               "DB919_ShotResultMach".ShotResult_Ma[1].Component.Comp[#Component].MaterialConsumption :=
               #TempConsumption +
               ("DB919_ShotResultMach".ShotResult_Ma[1].Component.Comp[#Component].Flow *
               "DB704_MH_Value".Mixinghead[#MHNumber].Corrvalue);

           ELSE
               "DB919_ShotResultMach".ShotResult_Ma[1].Component.Comp[#Component].MaterialConsumption :=
               #TempConsumption;

           END_IF;

       END_IF;
   END_FOR;
END_FUNCTION

ORGANIZATION_BLOCK "Cycle Execution"   // OB1, STL, ProgramCycle
TITLE = "Main Program Sweep (Cycle)"
{ S7_Optimized_Access := 'FALSE' }
VERSION : 0.1
   VAR_TEMP
      OB1_EV_CLASS : Byte;   // Bits 0-3 = 1 (Coming event), Bits 4-7 = 1 (Event class 1)
      OB1_SCAN_1 : Byte;   // 1 (Cold restart scan 1 of OB 1), 3 (Scan 2-n of OB 1)
      OB1_PRIORITY : Byte;   // Priority of OB Execution
      OB1_OB_NUMBR : Byte;   // 1 (Organization block 1, OB1)
      OB1_RESERVED_1 : Byte;   // Reserved for system
      OB1_RESERVED_2 : Byte;   // Reserved for system
      OB1_PREV_CYCLE : Int;   // Cycle time of previous OB1 scan (milliseconds)
      OB1_MIN_CYCLE : Int;   // Minimum cycle time of OB1 (milliseconds)
      OB1_MAX_CYCLE : Int;   // Maximum cycle time of OB1 (milliseconds)
      OB1_DATE_TIME : Date_And_Time;   // Date and time OB1 started
      Ret_Val_SFC51 : Int;
      SLZ_Header : Struct
         LENTHDR : Word;
         N_DR : Word;
      END_STRUCT;
      TmpMachineNo : Int;
      DPDPoff : Bool;
      RetValSFC : Int;
      DPDPon : Bool;
      D_ACT_DP_Busy : Bool;
   END_VAR
BEGIN

REGION Network 1: First PLC cycle
         A(;
         L     #OB1_SCAN_1;
         L     1;
         ==I;
         );
         =     "Flag_Erster_SPS_Zyklus";

   // --- Activate addresses of IO interface ProCan
         A     "Flag_Erster_SPS_Zyklus";
         S     "M1200_ActivateAdrProCan";
END_REGION

REGION Network 2: ProNet-Functions
         A     "Flag_Erster_SPS_Zyklus";
         R     "Flag_ToggleForDatarequest";

         CALL  "PNC_AI"
         ( RequestAll        := "Flag_Erster_SPS_Zyklus",
           AcknowledgeFaults := "DB009_Faults".Faults_Reset_FKT_M1,
           GOON              := "Flag_ToggleForDatarequest"
         );

         CALL  "PNC_Mixinghead"
         ( RequestAll        := "Flag_Erster_SPS_Zyklus",
           AcknowledgeFaults := "DB009_Faults".Faults_Reset_FKT_M1,
           GOON              := "Flag_ToggleForDatarequest"
         );

         CALL  "PNC_Flow"
         ( RequestAll        := "Flag_Erster_SPS_Zyklus",
           AcknowledgeFaults := "DB009_Faults".Faults_Reset_FKT_M1,
           GOON              := "Flag_ToggleForDatarequest"
         );

         AN    "Flag_ToggleForDatarequest";
         =     "Flag_ToggleForDatarequest";
END_REGION

REGION Network 3: Brücken für Inbetriebnahme
         CLR;
         =     "With_MC03";
         =     "With_MC04";
END_REGION

REGION Network 4: Handling Mould Editor
         CALL  "FB_MouldEditor_HMI", "FB_MouldEditor_HMI_DB"
         ( INiAmountMeteringUnits := "DB790_PlantParameter".AmountMeteringUnits,
           IOuMouldEditor_HMI     := "DB_MouldEditor_HMI".uData
         );
END_REGION

REGION Network 5: Analyse der Profinet- und Profibusbusteilnehmer
   // PN devices analyze
         CALL  DeviceStates
         ( LADDR   := "PN_Devices".LADDR,
           MODE    := "PN_Devices".MODE,
           Ret_Val := "PN_Devices".RETVAL,
           STATE   := "PN_Devices".Device_available
         );

   // PB devices analyze
         CALL  DeviceStates
         ( LADDR   := "PB_Devices".LADDR,
           MODE    := "PB_Devices".MODE,
           Ret_Val := "PB_Devices".RETVAL,
           STATE   := "PB_Devices".Device_available
         );
END_REGION

REGION Network 6: Tempering
   // Test
         CALL  "Baustein_1";

         O     "DB702_Tank_Value".Tank[1].With_Tempering_TempGeraet;
         O     "DB702_Tank_Value".Tank[1].With_Tempering_VKaltwasser;
         O     "DB702_Tank_Value".Tank[1].With_Tempering_Heizung;
         O     "DB702_Tank_Value".Tank[1].With_Tempering_WTRL;
         O     "DB702_Tank_Value".Tank[1].With_Tempering_WTmitFischer;
         O     "DB702_Tank_Value".Tank[1].With_Tempering_WTBypass;
         O     "DB702_Tank_Value".Tank[1].With_Tempering_WTVL;
   // Damit der Schalter für die Temperierung angezeigt wird
         =     "DB702_Tank_Value".Tank[1].With_Tempering;

         O     "DB702_Tank_Value".Tank[2].With_Tempering_TempGeraet;
         O     "DB702_Tank_Value".Tank[2].With_Tempering_VKaltwasser;
         O     "DB702_Tank_Value".Tank[2].With_Tempering_Heizung;
         O     "DB702_Tank_Value".Tank[2].With_Tempering_WTRL;
         O     "DB702_Tank_Value".Tank[2].With_Tempering_WTmitFischer;
         O     "DB702_Tank_Value".Tank[2].With_Tempering_WTBypass;
         O     "DB702_Tank_Value".Tank[2].With_Tempering_WTVL;
         =     "DB702_Tank_Value".Tank[2].With_Tempering;

         O     "DB702_Tank_Value".Tank[3].With_Tempering_TempGeraet;
         O     "DB702_Tank_Value".Tank[3].With_Tempering_VKaltwasser;
         O     "DB702_Tank_Value".Tank[3].With_Tempering_Heizung;
         O     "DB702_Tank_Value".Tank[3].With_Tempering_WTRL;
         O     "DB702_Tank_Value".Tank[3].With_Tempering_WTmitFischer;
         O     "DB702_Tank_Value".Tank[3].With_Tempering_WTBypass;
         O     "DB702_Tank_Value".Tank[3].With_Tempering_WTVL;
         =     "DB702_Tank_Value".Tank[3].With_Tempering;

         O     "DB702_Tank_Value".Tank[4].With_Tempering_TempGeraet;
         O     "DB702_Tank_Value".Tank[4].With_Tempering_VKaltwasser;
         O     "DB702_Tank_Value".Tank[4].With_Tempering_Heizung;
         O     "DB702_Tank_Value".Tank[4].With_Tempering_WTRL;
         O     "DB702_Tank_Value".Tank[4].With_Tempering_WTmitFischer;
         O     "DB702_Tank_Value".Tank[4].With_Tempering_WTBypass;
         O     "DB702_Tank_Value".Tank[4].With_Tempering_WTVL;
         =     "DB702_Tank_Value".Tank[4].With_Tempering;
END_REGION

REGION Network 7: Inputs external plant
   // MC1
   //      CALL  DPRD_DAT
   //         LADDR   :="PN-PN-Coupler_PU_MC1~IN___8_Byte"
   //         RET_VAL :=#RetValSFC
   //         RECORD  :="DB005_RS<->Extern".MC_Interface[1].Data_from_MC
   // MC2
   //     CALL  DPRD_DAT
   //         LADDR   :="PN-PN-Coupler_PU_MC2~IN__16_Byte"
   //         RET_VAL :=#RetValSFC
   //         RECORD  :="DB005_RS<->Extern".MC_Interface[2].Data_from_MC
   // MC3
   //      CALL  DPRD_DAT
   //         LADDR   :="PN-PN-Coupler_PU_MC3~IN__16_Byte"
   //         RET_VAL :=#RetValSFC
   //         RECORD  :="DB005_RS<->Extern".MC_Interface[3].Data_from_MC

   // MC4
   //      CALL  DPRD_DAT
   //         LADDR   :="PN-PN-Coupler_PU_MC4~IN__16_Byte"
   //         RET_VAL :=#RetValSFC
   //         RECORD  :="DB005_RS<->Extern".MC_Interface[4].Data_from_MC
END_REGION

REGION Network 8: Force Inputs
   //      L     "Interface_Signals_From_KMI":P
   //      T     %DB5.DBW20
   //      L     "Tag_35":P
   //      T     "DB005_RS<->Extern".MC_Interface[1].FromMC.Temperature_Tool01
   //      L     "Tag_36":P
   //      T     "DB005_RS<->Extern".MC_Interface[1].FromMC.Temperature_Tool02
   //      L     "Tag_37":P
   //      T     "DB005_RS<->Extern".MC_Interface[1].FromMC.Spare_6
   //      L     "Tag_38":P
   //      T     "DB005_RS<->Extern".MC_Interface[1].FromMC.Spare_8

   //      L     "Tag_39":P
   //      T     %DB5.DBW40
   //      L     "Tag_40":P
   //      T     "DB005_RS<->Extern".MC_Interface[2].FromMC.Temperature_Tool01
   //      L     "Tag_41":P
   //      T     "DB005_RS<->Extern".MC_Interface[2].FromMC.Temperature_Tool02
   //      L     "Tag_42":P
   //      T     "DB005_RS<->Extern".MC_Interface[2].FromMC.Spare_6
   //      L     "Tag_43":P
   //      T     "DB005_RS<->Extern".MC_Interface[2].FromMC.Spare_8
END_REGION

REGION Network 9: Check Profnet Slaves
   //
         CALL  DeviceStates
         ( LADDR   := 257,
           MODE    := 4,
           Ret_Val := #Ret_Val_SFC51,
           STATE   := "PN_DeviceState".StatePN
         );
   //
END_REGION

REGION Network 10: Interface Visu
         CALL  "FC5011_InterfaceHydraulik"
         ( Enable := 1
         );

         CALL  "FC5012_InterfaceTank"
         ( Enable := 1
         );

         CALL  "FC5013_InterfaceMetering"
         ( Enable := 1
         );

         CALL  "FC5014_InterfaceMixinghead"
         ( Enable := 1
         );

         CALL  "FC5020_InterfaceConfig"
         ( Enable := 1
         );

         CALL  "FC5900_InterfaceRobots"
         ( Enable := 1
         );
END_REGION

REGION Network 11: Program blocks
   //
         UC    "FB009_Faults";

   // machine 1
         UC    "FB011_OP_CirceMode_M1";
         UC    "FB012_MH_Hydraulic_M1";
         UC    "FB014_MH_SWU_M1";
         UC    "FB015_MeteringPump_M1";
   //     UC    "FB016_MeteringPump_Heating_M1"
         UC    "FB019_FoamingCycle_M1";
         UC    "FB017_CPiston_M1";

   // common function blocks
         UC    "FB100_Common_Aggregates_General";
         UC    "FB101_Common_Aggregates_C1";
         UC    "FB102_Common_Aggregates_C2";

         UC    "FB110_Interface_Prog_M1";
   //      UC    "FB111_Inerting"

         UC    "FB120_ProcanIO_RW";
   //      UC    "FB130_Tempering"
   //      UC    "FB140_ConfProCan"

         UC    "FB916_PV_LimitControl";

         UC    "FB919_PV_SetValueFoaming";
         UC    "FB920_ShotResult";

         UC    "FB930_FoamingData";

   //      UC    "FB1900_IF_Robots"

         UC    "FB1025_Service";

         CALL  "FC14_TP_Shortcuts";

   // Interface
         CALL  "FC2001_KM_FRA";
END_REGION

REGION Network 12: General functions
END_REGION

REGION Network 13: Outputs external plant
   // MC1
   //    CALL  DPWR_DAT
   //         LADDR   :="PN-PN-Coupler_PU_MC1~OUT___8_Byte"
   //         RECORD  :="DB005_RS<->Extern".MC_Interface[1].Data_to_MC
   //         RET_VAL :=#RetValSFC
   // MC2
   //     CALL  DPWR_DAT
   //         LADDR   :="PN-PN-Coupler_PU_MC2~OUT__16_Byte"
   //         RECORD  :="DB005_RS<->Extern".MC_Interface[2].Data_to_MC
   //         RET_VAL :=#RetValSFC
   // MC3
   //      CALL  DPWR_DAT
   //         LADDR   :="PN-PN-Coupler_PU_MC3~OUT__16_Byte"
   //         RECORD  :="DB005_RS<->Extern".MC_Interface[3].Data_to_MC
   //         RET_VAL :=#RetValSFC
   // MC4
   //      CALL  DPWR_DAT
   //         LADDR   :="PN-PN-Coupler_PU_MC4~OUT__16_Byte"
   //         RECORD  :="DB005_RS<->Extern".MC_Interface[4].Data_to_MC
   //         RET_VAL :=#RetValSFC
END_REGION

REGION Network 14: AllocationList
         CALL  "FB1931_ToolAllocationList", "FB1931_ToolAllocationList_DB";
END_REGION

REGION Network 15: Oszi
         CALL  "FC025_Oszilloskop";
         CALL  "FC117_INT_Umwandler";
END_REGION

REGION Network 16: TurnTable
   //    UC    "FB1001_TT"
END_REGION

REGION Network 17: RFID

   //      CALL  "FC030_BalluffReader 1"
   //      CALL  "FC031_BalluffReader 2"
END_REGION

REGION Network 18: Traceability
         CALL  "FC1500_ShotDataToMC";
END_REGION

REGION Network 19: Date and time
         CALL  "FC2170_TimeHandle";
   //-----
END_REGION

REGION Network 20: Network connection flag
         A     "Flag_00_500_Hertz";
         =     "Flag_Network";
END_REGION

REGION Network 21: delay_timer
         A     "new_shift";
         L     s5t#60s;
         SD    "delay_timer";
         A     "delay_timer";
         R     "new_shift";

         AN    "new_shift";
         R     "flag_delay_check_path";
         L     s5t#20s;
         SD    "Timer_check_path";
         A     "Timer_check_path";
         S     "flag_delay_check_path";
         R     "delay_timer";
END_REGION

REGION Network 22: IBN
         A     "AlwaysFALSE";
         R     "AlwaysFALSE";
         AN    "AlwaysTRUE";
         S     "AlwaysTRUE";
END_REGION
END_ORGANIZATION_BLOCK

ORGANIZATION_BLOCK "CYC_INT5"   // OB35, STL, CyclicInterrupt
TITLE = "Cyclic Interrupt"
{ S7_Optimized_Access := 'FALSE' }
AUTHOR : KT242
VERSION : 0.1
   VAR_TEMP
      OB35_EV_CLASS : Byte;   // Bits 0-3 = 1 (Coming event), Bits 4-7 = 1 (Event class 1)
      OB35_STRT_INF : Byte;   // 16#36 (OB 35 has started)
      OB35_PRIORITY : Byte;   // Priority of OB Execution
      OB35_OB_NUMBR : Byte;   // 35 (Organization block 35, OB35)
      OB35_RESERVED_1 : Byte;   // Reserved for system
      OB35_RESERVED_2 : Byte;   // Reserved for system
      OB35_PHASE_OFFSET : Word;   // Phase offset (msec)
      OB35_RESERVED_3 : Int;   // Reserved for system
      OB35_EXC_FREQ : Int;   // Frequency of execution (msec)
      OB35_DATE_TIME : Date_And_Time;   // Date and time OB35 started
      Temp_MH_Temp_C1 : Int;
      Temp_MH_Temp_C2 : Int;
      Temp_MH_Pressure_C1 : Int;
      Temp_MH_Pressure_C2 : Int;
      DINT_dummy : Real;
      dummy : Bool;
      Tenmp_flow_comp1 : DInt;
      Tenmp_flow_comp2 : DInt;
      Temp_ShotTimeAct : DInt;
      TempDBNo : Word;
      TempDWNo : DInt;
      TempRetClock : Int;
      TempDateTime : Date_And_Time;
      TempWritePointer : Int;
      EXC_FREQ_HE : Int;   // Execution frequency of heat exchangers
      TempSWU_MH01 : Bool;
      TempSWU_MH02 : Bool;
      TempSWU_MH03 : Bool;
      TempSWU_MH04 : Bool;
      TempSWU_MH05 : Bool;
      TempSWU_MH06 : Bool;
      TempSWU_MH07 : Bool;
      TempSWU_MH08 : Bool;
      TempSWU_MH09 : Bool;
      TempSWU_MH10 : Bool;
      Temp_CompFlowReal : Real;
      Temp_STimeReal : Real;
      CompUsedForShot : Array[1..16] of Bool;
   END_VAR
BEGIN

REGION Network 1: Read PV flowrate and calc. consumption of components machine 1
         A     "DB619_State_MPart".Cycle[1].Shotrelease;
         FP    "FHF_ShotreleaseM1";
         JCN   f101;
         L     0.0;
         T     "AmountFlowValuesMa1C1";
         T     "AmountFlowValuesMa1C2";
         T     "AmountFlowValuesMa1C3";
         T     "AmountFlowValuesMa1C4";
         T     "AmountFlowValuesMa1C5";
         T     "AmountFlowValuesMa1C6";
         T     "AmountFlowValuesMa1C7";
         T     "AmountFlowValuesMa1C8";
         T     "AmountFlowValuesMa1C9";
         T     "AmountFlowValuesMa1C10";
         T     "AmountFlowValuesMa1C11";
         T     "AmountFlowValuesMa1C12";

         T     "TotalFlowShotC01";
         T     "TotalFlowShotC02";
         T     "TotalFlowShotC03";
         T     "TotalFlowShotC04";
         T     "TotalFlowShotC05";
         T     "TotalFlowShotC06";
         T     "TotalFlowShotC07";
         T     "TotalFlowShotC08";
         T     "TotalFlowShotC09";
         T     "TotalFlowShotC10";
         T     "TotalFlowShotC11";
         T     "TotalFlowShotC12";


         T     "DB919_ShotResultMach".ShotResult_Ma[1].General.FoamingTime;
         T     "DB919_ShotResultMach".ShotResult_Ma[1].Component.Comp[1].Flow;
         T     "DB919_ShotResultMach".ShotResult_Ma[1].Component.Comp[2].Flow;
         T     "DB919_ShotResultMach".ShotResult_Ma[1].Component.Comp[3].Flow;
         T     "DB919_ShotResultMach".ShotResult_Ma[1].Component.Comp[4].Flow;
         T     "DB919_ShotResultMach".ShotResult_Ma[1].Component.Comp[5].Flow;
         T     "DB919_ShotResultMach".ShotResult_Ma[1].Component.Comp[6].Flow;
         T     "DB919_ShotResultMach".ShotResult_Ma[1].Component.Comp[7].Flow;
         T     "DB919_ShotResultMach".ShotResult_Ma[1].Component.Comp[8].Flow;
         T     "DB919_ShotResultMach".ShotResult_Ma[1].Component.Comp[9].Flow;
         T     "DB919_ShotResultMach".ShotResult_Ma[1].Component.Comp[10].Flow;
         T     "DB919_ShotResultMach".ShotResult_Ma[1].Component.Comp[11].Flow;
         T     "DB919_ShotResultMach".ShotResult_Ma[1].Component.Comp[12].Flow;


         T     "DB919_ShotResultMach".ShotResult_Ma[1].Component.Comp[1].MaterialConsumption;
         T     "DB919_ShotResultMach".ShotResult_Ma[1].Component.Comp[2].MaterialConsumption;
         T     "DB919_ShotResultMach".ShotResult_Ma[1].Component.Comp[3].MaterialConsumption;
         T     "DB919_ShotResultMach".ShotResult_Ma[1].Component.Comp[4].MaterialConsumption;
         T     "DB919_ShotResultMach".ShotResult_Ma[1].Component.Comp[5].MaterialConsumption;
         T     "DB919_ShotResultMach".ShotResult_Ma[1].Component.Comp[6].MaterialConsumption;
         T     "DB919_ShotResultMach".ShotResult_Ma[1].Component.Comp[7].MaterialConsumption;
         T     "DB919_ShotResultMach".ShotResult_Ma[1].Component.Comp[8].MaterialConsumption;
         T     "DB919_ShotResultMach".ShotResult_Ma[1].Component.Comp[9].MaterialConsumption;
         T     "DB919_ShotResultMach".ShotResult_Ma[1].Component.Comp[10].MaterialConsumption;
         T     "DB919_ShotResultMach".ShotResult_Ma[1].Component.Comp[11].MaterialConsumption;
         T     "DB919_ShotResultMach".ShotResult_Ma[1].Component.Comp[12].MaterialConsumption;

   //*******************************************************************************
   // ---- Flow COMPONENT 1 -----------------------
   f101: NOP   0;

         CALL  "FC920_PV_Calc_Act_Value"
         ( IN_Act_Value_read := "M1C01active",
           IN_Act_Value_ext  := FALSE,
           IN_Ext_Value      := #DINT_dummy,
           IN_Read_Double    := TRUE,
           IN_FLT_Needful    := 1,
           IN_FLT_Reset      := "DB009_Faults".HF_FaultsQuitOB35,
           IO_Any_ArrayPV    := "DB608_PV_Metering".Metering[1].Flow,
           IO_Fault_Sensor   := "DB823_Error_Metering".Flow_Component[1].Sensor_FLT_broken_wire,
           IO_New_Fault      := "DB009_Faults".Faultschanging_M1,
           IO_FLT_Level_3    := "DB009_Faults".Faults_FKT_Grp_3_M1
         );


   // --- Material consumption during shot component 1 ----
         ON    "M_ShotActive";  // "DB610_State_MPart".Cycle_Ma[1].ShotRuns
         ON    "M1C01active";
         JC    f102;
         A     "DB614_MH_State".MH_Status[1].Switch_Testshot_B_ON_OFF;
         L     0.0;
         JC    B1;
         L     "DB608_PV_Metering".Metering[1].Flow.PV_ActV.Value;
   B1:   L     "TotalFlowShotC01";
         +R;
         T     "TotalFlowShotC01";

         L     "AmountFlowValuesMa1C1";
         L     1.0;
         +R;
         T     "AmountFlowValuesMa1C1";

   //*******************************************************************************
   // ---- Flow COMPONENT 2 ---------------
   f102: NOP   0;

         CALL  "FC920_PV_Calc_Act_Value"
         ( IN_Act_Value_read := "M1C02active",
           IN_Act_Value_ext  := FALSE,
           IN_Ext_Value      := #DINT_dummy,
           IN_Read_Double    := TRUE,
           IN_FLT_Needful    := 1,
           IN_FLT_Reset      := "DB009_Faults".HF_FaultsQuitOB35,
           IO_Any_ArrayPV    := "DB608_PV_Metering".Metering[2].Flow,
           IO_Fault_Sensor   := "DB823_Error_Metering".Flow_Component[2].Sensor_FLT_broken_wire,
           IO_New_Fault      := "DB009_Faults".Faultschanging_M1,
           IO_FLT_Level_3    := "DB009_Faults".Faults_FKT_Grp_3_M1
         );


   // --- Material consumption during shot component 2 ---
         ON    "M_ShotActive";  // "DB610_State_MPart".Cycle_Ma[1].ShotRuns
         ON    "M1C02active";
         JC    f103;
         A     "DB614_MH_State".MH_Status[1].Switch_Testshot_A_ON_OFF;
         L     0.0;
         JC    B2;
         L     "DB608_PV_Metering".Metering[2].Flow.PV_ActV.Value;
   B2:   L     "TotalFlowShotC02";
         +R;
         T     "TotalFlowShotC02";

         L     "AmountFlowValuesMa1C2";
         L     1.0;
         +R;
         T     "AmountFlowValuesMa1C2";

   //*******************************************************************************
   // ---- Flow COMPONENT 3 ---------------
   f103: NOP   0;

         CALL  "FC920_PV_Calc_Act_Value"
         ( IN_Act_Value_read := "M1C03active",
           IN_Act_Value_ext  := FALSE,
           IN_Ext_Value      := #DINT_dummy,
           IN_Read_Double    := TRUE,
           IN_FLT_Needful    := 1,
           IN_FLT_Reset      := "DB009_Faults".HF_FaultsQuitOB35,
           IO_Any_ArrayPV    := "DB608_PV_Metering".Metering[3].Flow,
           IO_Fault_Sensor   := "DB823_Error_Metering".Flow_Component[3].Sensor_FLT_broken_wire,
           IO_New_Fault      := "DB009_Faults".Faultschanging_M1,
           IO_FLT_Level_3    := "DB009_Faults".Faults_FKT_Grp_3_M1
         );


   // --- Material consumption during shot component 3 ---
         ON    "M_ShotActive";  // "DB610_State_MPart".Cycle_Ma[1].ShotRuns
         ON    "M1C03active";
         JC    f104;
         L     "DB608_PV_Metering".Metering[3].Flow.PV_ActV.Value;
         L     "TotalFlowShotC03";
         +R;
         T     "TotalFlowShotC03";

         L     "AmountFlowValuesMa1C3";
         L     1.0;
         +R;
         T     "AmountFlowValuesMa1C3";

   //*******************************************************************************
   // ---- Flow COMPONENT 4 ---------------
   f104: NOP   0;

         CALL  "FC920_PV_Calc_Act_Value"
         ( IN_Act_Value_read := "M1C04active",
           IN_Act_Value_ext  := FALSE,
           IN_Ext_Value      := #DINT_dummy,
           IN_Read_Double    := TRUE,
           IN_FLT_Needful    := 1,
           IN_FLT_Reset      := "DB009_Faults".HF_FaultsQuitOB35,
           IO_Any_ArrayPV    := "DB608_PV_Metering".Metering[4].Flow,
           IO_Fault_Sensor   := "DB823_Error_Metering".Flow_Component[4].Sensor_FLT_broken_wire,
           IO_New_Fault      := "DB009_Faults".Faultschanging_M1,
           IO_FLT_Level_3    := "DB009_Faults".Faults_FKT_Grp_3_M1
         );


   // --- Material consumption during shot component 4 ---
         ON    "M_ShotActive";  // "DB610_State_MPart".Cycle_Ma[1].ShotRuns
         ON    "M1C04active";
         JC    f105;
         L     "DB608_PV_Metering".Metering[4].Flow.PV_ActV.Value;
         L     "TotalFlowShotC04";
         +R;
         T     "TotalFlowShotC04";

         L     "AmountFlowValuesMa1C4";
         L     1.0;
         +R;
         T     "AmountFlowValuesMa1C4";

   //*******************************************************************************
   // ---- Flow COMPONENT 5 ---------------
   f105: NOP   0;

         CALL  "FC920_PV_Calc_Act_Value"
         ( IN_Act_Value_read := "M1C05active",
           IN_Act_Value_ext  := FALSE,
           IN_Ext_Value      := #DINT_dummy,
           IN_Read_Double    := TRUE,
           IN_FLT_Needful    := 1,
           IN_FLT_Reset      := "DB009_Faults".HF_FaultsQuitOB35,
           IO_Any_ArrayPV    := "DB608_PV_Metering".Metering[5].Flow,
           IO_Fault_Sensor   := "DB823_Error_Metering".Flow_Component[5].Sensor_FLT_broken_wire,
           IO_New_Fault      := "DB009_Faults".Faultschanging_M1,
           IO_FLT_Level_3    := "DB009_Faults".Faults_FKT_Grp_3_M1
         );


   // --- Material consumption during shot component 5 ---
         ON    "M_ShotActive";  // "DB610_State_MPart".Cycle_Ma[1].ShotRuns
         ON    "M1C05active";
         JC    f106;
         L     "DB608_PV_Metering".Metering[5].Flow.PV_ActV.Value;
         L     "TotalFlowShotC05";
         +R;
         T     "TotalFlowShotC05";

         L     "AmountFlowValuesMa1C5";
         L     1.0;
         +R;
         T     "AmountFlowValuesMa1C5";

   //*******************************************************************************
   // ---- Flow COMPONENT 6 ---------------
   f106: NOP   0;

         CALL  "FC920_PV_Calc_Act_Value"
         ( IN_Act_Value_read := "M1C06active",
           IN_Act_Value_ext  := FALSE,
           IN_Ext_Value      := #DINT_dummy,
           IN_Read_Double    := TRUE,
           IN_FLT_Needful    := 1,
           IN_FLT_Reset      := "DB009_Faults".HF_FaultsQuitOB35,
           IO_Any_ArrayPV    := "DB608_PV_Metering".Metering[6].Flow,
           IO_Fault_Sensor   := "DB823_Error_Metering".Flow_Component[6].Sensor_FLT_broken_wire,
           IO_New_Fault      := "DB009_Faults".Faultschanging_M1,
           IO_FLT_Level_3    := "DB009_Faults".Faults_FKT_Grp_3_M1
         );


   // --- Material consumption during shot component 6 ---
         ON    "M_ShotActive";  // "DB610_State_MPart".Cycle_Ma[1].ShotRuns
         ON    "M1C06active";
         JC    f107;
         L     "DB608_PV_Metering".Metering[6].Flow.PV_ActV.Value;
         L     "TotalFlowShotC06";
         +R;
         T     "TotalFlowShotC06";

         L     "AmountFlowValuesMa1C6";
         L     1.0;
         +R;
         T     "AmountFlowValuesMa1C6";

   //*******************************************************************************
   // ---- Flow COMPONENT 7 ---------------
   f107: NOP   0;

         CALL  "FC920_PV_Calc_Act_Value"
         ( IN_Act_Value_read := "M1C07active",
           IN_Act_Value_ext  := FALSE,
           IN_Ext_Value      := #DINT_dummy,
           IN_Read_Double    := TRUE,
           IN_FLT_Needful    := 1,
           IN_FLT_Reset      := "DB009_Faults".HF_FaultsQuitOB35,
           IO_Any_ArrayPV    := "DB608_PV_Metering".Metering[7].Flow,
           IO_Fault_Sensor   := "DB823_Error_Metering".Flow_Component[7].Sensor_FLT_broken_wire,
           IO_New_Fault      := "DB009_Faults".Faultschanging_M1,
           IO_FLT_Level_3    := "DB009_Faults".Faults_FKT_Grp_3_M1
         );


   // --- Material consumption during shot component 7 ---
         ON    "M_ShotActive";  // "DB610_State_MPart".Cycle_Ma[1].ShotRuns
         ON    "M1C07active";
         JC    f108;
         L     "DB608_PV_Metering".Metering[7].Flow.PV_ActV.Value;
         L     "TotalFlowShotC07";
         +R;
         T     "TotalFlowShotC07";

         L     "AmountFlowValuesMa1C7";
         L     1.0;
         +R;
         T     "AmountFlowValuesMa1C7";

   //*******************************************************************************
   // ---- Flow COMPONENT 8 ---------------
   f108: NOP   0;

         CALL  "FC920_PV_Calc_Act_Value"
         ( IN_Act_Value_read := "M1C08active",
           IN_Act_Value_ext  := FALSE,
           IN_Ext_Value      := #DINT_dummy,
           IN_Read_Double    := TRUE,
           IN_FLT_Needful    := 1,
           IN_FLT_Reset      := "DB009_Faults".HF_FaultsQuitOB35,
           IO_Any_ArrayPV    := "DB608_PV_Metering".Metering[8].Flow,
           IO_Fault_Sensor   := "DB823_Error_Metering".Flow_Component[8].Sensor_FLT_broken_wire,
           IO_New_Fault      := "DB009_Faults".Faultschanging_M1,
           IO_FLT_Level_3    := "DB009_Faults".Faults_FKT_Grp_3_M1
         );


   // --- Material consumption during shot component 8 ---
         ON    "M_ShotActive";  // "DB610_State_MPart".Cycle_Ma[1].ShotRuns
         ON    "M1C08active";
         JC    f109;
         L     "DB608_PV_Metering".Metering[8].Flow.PV_ActV.Value;
         L     "TotalFlowShotC08";
         +R;
         T     "TotalFlowShotC08";

         L     "AmountFlowValuesMa1C8";
         L     1.0;
         +R;
         T     "AmountFlowValuesMa1C8";

   //*******************************************************************************
   // ---- Flow COMPONENT 9 ---------------
   f109: NOP   0;

         CALL  "FC920_PV_Calc_Act_Value"
         ( IN_Act_Value_read := "M1C09active",
           IN_Act_Value_ext  := FALSE,
           IN_Ext_Value      := #DINT_dummy,
           IN_Read_Double    := TRUE,
           IN_FLT_Needful    := 1,
           IN_FLT_Reset      := "DB009_Faults".HF_FaultsQuitOB35,
           IO_Any_ArrayPV    := "DB608_PV_Metering".Metering[09].Flow,
           IO_Fault_Sensor   := "DB823_Error_Metering".Flow_Component[09].Sensor_FLT_broken_wire,
           IO_New_Fault      := "DB009_Faults".Faultschanging_M1,
           IO_FLT_Level_3    := "DB009_Faults".Faults_FKT_Grp_3_M1
         );


   // --- Material consumption during shot component 09 ---
         ON    "M_ShotActive";  // "DB610_State_MPart".Cycle_Ma[1].ShotRuns
         ON    "M1C09active";
         JC    f110;
         L     "DB608_PV_Metering".Metering[9].Flow.PV_ActV.Value;
         L     "TotalFlowShotC09";
         +R;
         T     "TotalFlowShotC09";

         L     "AmountFlowValuesMa1C9";
         L     1.0;
         +R;
         T     "AmountFlowValuesMa1C9";

   //*******************************************************************************
   // ---- Flow COMPONENT 10 ---------------
   f110: NOP   0;

         CALL  "FC920_PV_Calc_Act_Value"
         ( IN_Act_Value_read := "M1C10active",
           IN_Act_Value_ext  := FALSE,
           IN_Ext_Value      := #DINT_dummy,
           IN_Read_Double    := TRUE,
           IN_FLT_Needful    := 1,
           IN_FLT_Reset      := "DB009_Faults".HF_FaultsQuitOB35,
           IO_Any_ArrayPV    := "DB608_PV_Metering".Metering[10].Flow,
           IO_Fault_Sensor   := "DB823_Error_Metering".Flow_Component[10].Sensor_FLT_broken_wire,
           IO_New_Fault      := "DB009_Faults".Faultschanging_M1,
           IO_FLT_Level_3    := "DB009_Faults".Faults_FKT_Grp_3_M1
         );


   // --- Material consumption during shot component 10 ---
         ON    "M_ShotActive";  // "DB610_State_MPart".Cycle_Ma[1].ShotRuns
         ON    "M1C10active";
         JC    f111;
         L     "DB608_PV_Metering".Metering[10].Flow.PV_ActV.Value;
         L     "TotalFlowShotC10";
         +R;
         T     "TotalFlowShotC10";

         L     "AmountFlowValuesMa1C10";
         L     1.0;
         +R;
         T     "AmountFlowValuesMa1C10";

   //*******************************************************************************
   // ---- Flow COMPONENT 11 ---------------
   f111: NOP   0;

         CALL  "FC920_PV_Calc_Act_Value"
         ( IN_Act_Value_read := "M1C11active",
           IN_Act_Value_ext  := FALSE,
           IN_Ext_Value      := #DINT_dummy,
           IN_Read_Double    := TRUE,
           IN_FLT_Needful    := 1,
           IN_FLT_Reset      := "DB009_Faults".HF_FaultsQuitOB35,
           IO_Any_ArrayPV    := "DB608_PV_Metering".Metering[11].Flow,
           IO_Fault_Sensor   := "DB823_Error_Metering".Flow_Component[11].Sensor_FLT_broken_wire,
           IO_New_Fault      := "DB009_Faults".Faultschanging_M1,
           IO_FLT_Level_3    := "DB009_Faults".Faults_FKT_Grp_3_M1
         );


   // --- Material consumption during shot component 11 ---
         ON    "M_ShotActive";  // "DB610_State_MPart".Cycle_Ma[1].ShotRuns
         ON    "M1C11active";
         JC    f112;
         L     "DB608_PV_Metering".Metering[11].Flow.PV_ActV.Value;
         L     "TotalFlowShotC11";
         +R;
         T     "TotalFlowShotC11";

         L     "AmountFlowValuesMa1C11";
         L     1.0;
         +R;
         T     "AmountFlowValuesMa1C11";

   //*******************************************************************************
   // ---- Flow COMPONENT 12 ---------------
   f112: NOP   0;

         CALL  "FC920_PV_Calc_Act_Value"
         ( IN_Act_Value_read := "M1C12active",
           IN_Act_Value_ext  := FALSE,
           IN_Ext_Value      := #DINT_dummy,
           IN_Read_Double    := TRUE,
           IN_FLT_Needful    := 1,
           IN_FLT_Reset      := "DB009_Faults".HF_FaultsQuitOB35,
           IO_Any_ArrayPV    := "DB608_PV_Metering".Metering[12].Flow,
           IO_Fault_Sensor   := "DB823_Error_Metering".Flow_Component[12].Sensor_FLT_broken_wire,
           IO_New_Fault      := "DB009_Faults".Faultschanging_M1,
           IO_FLT_Level_3    := "DB009_Faults".Faults_FKT_Grp_3_M1
         );


   // --- Material consumption during shot component 12 ---
         ON    "M_ShotActive";  // "DB610_State_MPart".Cycle_Ma[1].ShotRuns
         ON    "M1C12active";
         JC    f113;
         L     "DB608_PV_Metering".Metering[12].Flow.PV_ActV.Value;
         L     "TotalFlowShotC12";
         +R;
         T     "TotalFlowShotC12";

         L     "AmountFlowValuesMa1C12";
         L     1.0;
         +R;
         T     "AmountFlowValuesMa1C12";

   //*******************************************************************************
   // ---- Flow COMPONENT 13 ---------------
   f113: NOP   0;
   //*******************************************************************************
END_REGION

REGION Network 2: Read PV flowrate and calc. consumption of components machine 2
END_REGION

REGION Network 3: Shotdata: Shottime, Consumption of machine 1

         L     "TotalFlowShotC01";
         T     "DB919_ShotResultMach".TotalFlowShotM1[1];
         L     "TotalFlowShotC02";
         T     "DB919_ShotResultMach".TotalFlowShotM1[2];
         L     "TotalFlowShotC03";
         T     "DB919_ShotResultMach".TotalFlowShotM1[3];
         L     "TotalFlowShotC04";
         T     "DB919_ShotResultMach".TotalFlowShotM1[4];
         L     "TotalFlowShotC05";
         T     "DB919_ShotResultMach".TotalFlowShotM1[5];
         L     "TotalFlowShotC06";
         T     "DB919_ShotResultMach".TotalFlowShotM1[6];
         L     "TotalFlowShotC07";
         T     "DB919_ShotResultMach".TotalFlowShotM1[7];
         L     "TotalFlowShotC08";
         T     "DB919_ShotResultMach".TotalFlowShotM1[8];
         L     "TotalFlowShotC09";
         T     "DB919_ShotResultMach".TotalFlowShotM1[9];
         L     "TotalFlowShotC10";
         T     "DB919_ShotResultMach".TotalFlowShotM1[10];
         L     "TotalFlowShotC11";
         T     "DB919_ShotResultMach".TotalFlowShotM1[11];
         L     "TotalFlowShotC12";
         T     "DB919_ShotResultMach".TotalFlowShotM1[12];

         L     "AmountFlowValuesMa1C1";
         T     "DB919_ShotResultMach".AmountFlowValuesM1[1];
         L     "AmountFlowValuesMa1C2";
         T     "DB919_ShotResultMach".AmountFlowValuesM1[2];
         L     "AmountFlowValuesMa1C3";
         T     "DB919_ShotResultMach".AmountFlowValuesM1[3];
         L     "AmountFlowValuesMa1C4";
         T     "DB919_ShotResultMach".AmountFlowValuesM1[4];
         L     "AmountFlowValuesMa1C5";
         T     "DB919_ShotResultMach".AmountFlowValuesM1[5];
         L     "AmountFlowValuesMa1C6";
         T     "DB919_ShotResultMach".AmountFlowValuesM1[6];
         L     "AmountFlowValuesMa1C7";
         T     "DB919_ShotResultMach".AmountFlowValuesM1[7];
         L     "AmountFlowValuesMa1C8";
         T     "DB919_ShotResultMach".AmountFlowValuesM1[8];
         L     "AmountFlowValuesMa1C9";
         T     "DB919_ShotResultMach".AmountFlowValuesM1[9];
         L     "AmountFlowValuesMa1C10";
         T     "DB919_ShotResultMach".AmountFlowValuesM1[10];
         L     "AmountFlowValuesMa1C11";
         T     "DB919_ShotResultMach".AmountFlowValuesM1[11];
         L     "AmountFlowValuesMa1C12";
         T     "DB919_ShotResultMach".AmountFlowValuesM1[12];


         A     "DB619_State_MPart".Cycle[1].ShotRuns;
         FP    "HF_FP_ShotRuns";
         JCN   n12s;
         L     "DB619_State_MPart".ShotMa[1].ShotData.Comp_at_Shot;
         T     "CompAtShot";

   n12s: A     "ShotStoppedM1";  // "DB610_State_MPart".Cycle_Ma[1].PulsShotend
         FP    "HF_FP_ShotStoppedM1";
         JCN   st1E;
         S     "CalcShotValuesMa1";

   // Copy Control bits for module to local area
         L;
         LAR1;
         L     "CompAtShot";
         CAW;
         T     LW[AR1, P#0.0];

         CALL  "ShotData_OB35"
         ( CompForShot := #CompUsedForShot
         );

   st1E: NOP   0;
END_REGION

REGION Network 4: Read prepressure of pumps
   // C1 M1
         CALL  "FC920_PV_Calc_Act_Value"
         ( IN_Act_Value_read := TRUE,
           IN_Act_Value_ext  := FALSE,
           IN_Ext_Value      := #DINT_dummy,
           IN_Read_Double    := FALSE,
           IN_FLT_Needful    := FALSE,
           IN_FLT_Reset      := "DB009_Faults".HF_FaultsQuitOB35,
           IO_Any_ArrayPV    := "DB608_PV_Metering".Metering[1].Pre_Pressure,
           IO_Fault_Sensor   := #dummy,
           IO_New_Fault      := "DB009_Faults".Faultschanging_M1,
           IO_FLT_Level_3    := "DB009_Faults".Faults_FKT_Grp_3_M1
         );

   // C2 M1
         CALL  "FC920_PV_Calc_Act_Value"
         ( IN_Act_Value_read := TRUE,
           IN_Act_Value_ext  := FALSE,
           IN_Ext_Value      := #DINT_dummy,
           IN_Read_Double    := FALSE,
           IN_FLT_Needful    := FALSE,
           IN_FLT_Reset      := "DB009_Faults".HF_FaultsQuitOB35,
           IO_Any_ArrayPV    := "DB608_PV_Metering".Metering[2].Pre_Pressure,
           IO_Fault_Sensor   := #dummy,
           IO_New_Fault      := "DB009_Faults".Faultschanging_M1,
           IO_FLT_Level_3    := "DB009_Faults".Faults_FKT_Grp_3_M1
         );
END_REGION

REGION Network 5: Read flow of pneumatics unit
         CALL  "FC920_PV_Calc_Act_Value"
         ( IN_Act_Value_read := TRUE,
           IN_Act_Value_ext  := FALSE,
           IN_Ext_Value      := #DINT_dummy,
           IN_Read_Double    := FALSE,
           IN_FLT_Needful    := FALSE,
           IN_FLT_Reset      := "DB009_Faults".HF_FaultsQuitOB35,
           IO_Any_ArrayPV    := "DB606_PV_Machine".Machine[1].PneumaticFlow,
           IO_Fault_Sensor   := #dummy,
           IO_New_Fault      := "DB009_Faults".Faultschanging_M1,
           IO_FLT_Level_3    := "DB009_Faults".Faults_FKT_Grp_3_M1
         );
END_REGION

REGION Network 6: PID-control of prepressure
   // C1 M1
   //      CALL  "FC109_PID_FeedingPump"
   //         OB35_EXC_FREQ        :=#OB35_EXC_FREQ
   //         PID_ProportionalGain :="DB751_auxiliaryDriveMetering".FeedingPumpControler[1].ProportionalGain
   //         PID_ResetTime        :="DB751_auxiliaryDriveMetering".FeedingPumpControler[1].ResetTime
   //         PID_DerivativeTime   :="DB751_auxiliaryDriveMetering".FeedingPumpControler[1].DerivativeTime
   //         MaxValPAW            :=10000.0 //2.764800e+004
   //         ControllerOn         :="M_FeedingP_Start_C1"
   //         ByteSwapOutPut       :=FALSE
   //         Enable               :=TRUE
   //         FaultSensor          :=FALSE
   //         PAW                  :="Set_FeedingP_C1":P
   //         ManipValue_mV        :="DB613_Komponent_State".FeedPump[1].ManipValuePercent
   //         IO_PV                :="DB608_PV_Metering".Metering[1].Pre_Pressure
   //         IO_PIDStatus         :="DB613_Komponent_State".FeedingPumpControler[1]
   //         IO_PIDContrStatus    :="DB613_Komponent_State".FeedPump[1].State_Drive

   // C2 M1
   //      CALL  "FC109_PID_FeedingPump"
   //         OB35_EXC_FREQ        :=#OB35_EXC_FREQ
   //         PID_ProportionalGain :="DB751_auxiliaryDriveMetering".FeedingPumpControler[2].ProportionalGain
   //         PID_ResetTime        :="DB751_auxiliaryDriveMetering".FeedingPumpControler[2].ResetTime
   //         PID_DerivativeTime   :="DB751_auxiliaryDriveMetering".FeedingPumpControler[2].DerivativeTime
   //         MaxValPAW            :=10000.0 //2.764800e+004
   //         ControllerOn         :="M_FeedingP_Start_C2"
   //         ByteSwapOutPut       :=FALSE
   //         Enable               :=TRUE
   //         FaultSensor          :=FALSE
   //         PAW                  :="Set_FeedingP_C2":P
   //         ManipValue_mV        :="DB613_Komponent_State".FeedPump[2].ManipValuePercent
   //         IO_PV                :="DB608_PV_Metering".Metering[2].Pre_Pressure
   //         IO_PIDStatus         :="DB613_Komponent_State".FeedingPumpControler[2]
   //         IO_PIDContrStatus    :="DB613_Komponent_State".FeedPump[2].State_Drive
END_REGION

REGION Network 7: Shotdata: Shottime, Consumption of machine 2
END_REGION

REGION Network 8: Data sampling of oszi function
END_REGION

REGION Network 9: Measuring Inerting MH1
         A     "DB614_MH_State".InertingMH[1].Inert_runs;
         FP    "DB614_MH_State".InertingMH[1].FP_Start_Inert;
         =     "DB614_MH_State".InertingMH[1].FH_Start_Inert;

         ON    "DB614_MH_State".InertingMH[1].FP_Start_Inert;
         O     "DB614_MH_State".InertingMH[1].FH_Start_Inert;
         JC    weit;

         L     "DB614_MH_State".InertingMH[1].Actual_Flow_N2;
         L     "DB614_MH_State".InertingMH[1].Actual_Flow_N2_measured_Total;
         +R;
         T     "DB614_MH_State".InertingMH[1].Actual_Flow_N2_measured_Total;
         L     600.0;
         /R;
         T     "DB614_MH_State".InertingMH[1].Total_Flow_N2_Visu;
         JU    ende;

   weit: AN    "DB614_MH_State".InertingMH[1].FH_Start_Inert;
         JC    ende;
         L     0.0;
         T     "DB614_MH_State".InertingMH[1].Actual_Flow_N2_measured_Total;
         T     "DB614_MH_State".InertingMH[1].Total_Flow_N2_Visu;

   ende: L     "DB614_MH_State".InertingMH[1].Actual_Flow_N2;
         L     6.0;
         /R;
         T     "DB614_MH_State".InertingMH[1].Actual_Flow_N2_Visu;
END_REGION

REGION Network 10: Leakage measuring MH1
         A     "DB614_MH_State".InertingMH[1].Set_LoadValue;
         O     "V_Inert_Piston_MH1";
         O(;
         L     "DB704_MH_Value".MH_Inerting[1].Leakage_Value;
         L     0.0;
         ==D;
         );
         JC    Null;

         A     "T_Leakage_Ctrl_Tact_N2";
         FP    "DB614_MH_State".InertingMH[1].FP_Start_Leakage_Control;
         =     "DB614_MH_State".InertingMH[1].FH_Start_Leakage_Control;

         ON    "DB614_MH_State".InertingMH[1].FP_Start_Leakage_Control;
         O     "DB614_MH_State".InertingMH[1].FH_Start_Leakage_Control;
         JC    WLeak;

         L     "DB604_PV_Mixinghead".Mixinghead[1].Inerting.PV_ActV.Value;
         T     "DB614_MH_State".InertingMH[1].Actual_Flow_N2;

         L     "DB614_MH_State".InertingMH[1].Actual_Flow_N2;
         L     "DB614_MH_State".InertingMH[1].Leakage_Actual_Flow_N2_measured_Total;
         +R;
         T     "DB614_MH_State".InertingMH[1].Leakage_Actual_Flow_N2_measured_Total;
         L     600.0;
         /R;
         T     "DB614_MH_State".InertingMH[1].Leakage_Total_Flow_N2_Visu;
         JU    ELEAK;

   WLeak:AN    "DB614_MH_State".InertingMH[1].FH_Start_Leakage_Control;
         JC    ELEAK;
   Null: L     0.0;
         T     "DB614_MH_State".InertingMH[1].Leakage_Actual_Flow_N2_measured_Total;
         T     "DB614_MH_State".InertingMH[1].Leakage_Total_Flow_N2_Visu;
         SET;
         R     "DB614_MH_State".InertingMH[1].Set_LoadValue;
   ELEAK:L     "DB614_MH_State".InertingMH[1].Leakage_Total_Flow_N2_Visu;
         L     60.0;
         /R;
         T     "DB614_MH_State".InertingMH[1].Leakage_Actual_Flow_N2_Visu;
END_REGION

REGION Network 11: Reset HF_FaultsQuitOB35
         SET;
         R     "DB009_Faults".HF_FaultsQuitOB35;
END_REGION
END_ORGANIZATION_BLOCK

ORGANIZATION_BLOCK "CYCL_FLT"   // OB80, STL, TimeErrorInterrupt
TITLE = "Cycle Time Fault"
{ S7_Optimized_Access := 'FALSE' }
AUTHOR : KT242
VERSION : 0.0
   VAR_TEMP
      OB80_EV_CLASS : Byte;   // 16#35, Event class 3, Entering event state, Internal fault event
      OB80_FLT_ID : Byte;   // 16#XX, Fault identifcation code
      OB80_PRIORITY : Byte;   // Priority of OB Execution
      OB80_OB_NUMBR : Byte;   // 80 (Organization block 80, OB80)
      OB80_RESERVED_1 : Byte;   // Reserved for system
      OB80_RESERVED_2 : Byte;   // Reserved for system
      OB80_ERROR_INFO : Word;   // Error information on event
      OB80_ERR_EV_CLASS : Byte;   // Class of event causing error
      OB80_ERR_EV_NUM : Byte;   // Number of event causing error
      OB80_OB_PRIORITY : Byte;   // Priority of OB causing error
      OB80_OB_NUM : Byte;   // Number of OB causing error
      OB80_DATE_TIME : Date_And_Time;   // Date and time OB80 started
   END_VAR
BEGIN
END_ORGANIZATION_BLOCK

ORGANIZATION_BLOCK "Pull or plug of modules"   // OB83, LAD, PullPlug
{ S7_Optimized_Access := 'TRUE' }
VERSION : 0.1
   VAR_INPUT
      LADDR : Hw_Io;   // Hardware identifier
      Event_Class : Byte;   // 16#38/39: module inserted, removed
      Fault_ID : Byte;   // Fault identifier
   END_VAR
BEGIN
END_ORGANIZATION_BLOCK

ORGANIZATION_BLOCK "OB100_ANLAUF"   // OB100, STL, Startup
TITLE = Start up / new start
{ S7_Optimized_Access := 'FALSE' }
AUTHOR : KT242
VERSION : 0.1
   VAR_TEMP
      OB100_EV_CLASS : Byte;   // 16#13, Event class 1, Entering event state, Event logged in diagnostic buffer
      OB100_STRTUP : Byte;   // 16#81/82/83/84 Method of startup
      OB100_PRIORITY : Byte;   // 27 (Priority of 1 is lowest)
      OB100_OB_NUMBR : Byte;   // 100 (Organization block 100, OB100)
      OB100_RESERVED_1 : Byte;   // Reserved for system
      OB100_RESERVED_2 : Byte;   // Reserved for system
      OB100_STOP : Word;   // Event that caused CPU to stop (16#4xxx)
      OB100_STRT_INFO : DWord;   // Information on how system started
      OB100_DATE_TIME : Date_And_Time;   // Date and time OB100 started
      Ret_Val : Int;
   END_VAR
BEGIN

REGION Network 1: Request write values
END_REGION
END_ORGANIZATION_BLOCK

(* ===== HMI "HMI_RT_1" =====
system functions are stored by id; their names below are inferred from use
connection "HMI_Connection_2": ETHERNET, S7_1500_OMS

HMI tags "Default tag table"
   "NavUserChange" : Int, internal
   "NavScreenChange" : Int, internal
   "Alarm_Filter_Tag" : Int, internal
   "tes_1" : Bool, internal
   "tes_2" : Bool, internal
   "tes_3" : Bool, internal
   "Date_1" : DateTime, internal
   "Date" : DateTime, internal
   "Time" : DateTime, internal
   "HMI_Tag_1" : Int, internal
   "HMI_Tag_1(1)" : Int, internal
   "tes_Time_1" : DateTime, internal
   "tes_Time_2" : DateTime, internal
   "tes_Time_3" : DateTime, internal
   "L_DT_max_C1" : Bool = PLC DB14_TP_Shortcuts.TP_Shortcuts.ButtonNo.1 AT %I21.5, 1 s
   "L_Tank_min_C1" : Bool = PLC DB14_TP_Shortcuts.TP_Shortcuts.ButtonNo.2 AT %I21.2, 1 s
   "L_Tank_min_C2" : Bool = PLC DB14_TP_Shortcuts.TP_Shortcuts.ButtonNo.3 AT %I23.2, 1 s
   "L_DT_max_C2" : Bool = PLC DB14_TP_Shortcuts.TP_Shortcuts.ButtonNo.5 AT %I23.5, 1 s
   "PopUp_Restrict" : Bool, internal
   "return_result" : Int, internal

HMI tags "Machine"
   "DB619_State_MPart_Write" : Bool = PLC DB14_TP_Shortcuts.TP_Shortcuts.ButtonNo.5 AT %DB619.DBX6.1, 1 s
   "DB700_Machine_Machine{0}_CtrlChangeTime1" : S5Time = PLC DB14_TP_Shortcuts.TP_Shortcuts.Page_active.1 AT %DB700.DBW26, 1 s
      on ChangeValue: SetBit("DB619_State_MPart_Write")
   "DB700_Machine_Machine{0}_HP_time_after_shot" : S5Time = PLC DB14_TP_Shortcuts.TP_Shortcuts.Page_active.2 AT %DB700.DBW18, 1 s
      on ChangeValue: SetBit("DB619_State_MPart_Write")
   "DB700_Machine_Machine{0}_Int_Pausetime_Auto" : S5Time = PLC DB14_TP_Shortcuts.TP_Shortcuts.ButtonNo.2 AT %DB700.DBW12, 1 s
      on ChangeValue: SetBit("DB619_State_MPart_Write")
   "DB700_Machine_Machine{0}_Int_Pausetime_Manual" : S5Time = PLC DB14_TP_Shortcuts.TP_Shortcuts.ButtonNo.7 AT %DB700.DBW8, 1 s
      on ChangeValue: SetBit("DB619_State_MPart_Write")
   "DB700_Machine_Machine{0}_Int_Runtime_Auto" : S5Time = PLC DB14_TP_Shortcuts.TP_Shortcuts.ButtonNo.1 AT %DB700.DBW10, 1 s
      on ChangeValue: SetBit("DB619_State_MPart_Write")
   "DB700_Machine_Machine{0}_Int_Runtime_Manual" : S5Time = PLC DB14_TP_Shortcuts.TP_Shortcuts.ButtonNo.3 AT %DB700.DBW6, 1 s
      on ChangeValue: SetBit("DB619_State_MPart_Write")
   "DB700_Machine_Machine{0}_Max_ShotTime" : S5Time = PLC DB14_TP_Shortcuts.TP_Shortcuts.Page_active.4 AT %DB700.DBW30, 1 s
      on ChangeValue: SetBit("DB619_State_MPart_Write")
   "DB700_Machine_Machine{0}_Max_WaitTime" : S5Time = PLC DB14_TP_Shortcuts.TP_Shortcuts.Page_active.5 AT %DB700.DBW34, 1 s
      on ChangeValue: SetBit("DB619_State_MPart_Write")
   "DB700_Machine_Machine{0}_Min_ShotTime" : S5Time = PLC DB14_TP_Shortcuts.TP_Shortcuts.Page_active.3 AT %DB700.DBW32, 1 s
      on ChangeValue: SetBit("DB619_State_MPart_Write")
   "DB700_Machine_Machine{0}_PressureBuildUpTime" : S5Time = PLC DB14_TP_Shortcuts.TP_Shortcuts.Page_active.6 AT %DB700.DBW22, 1 s
      on ChangeValue: SetBit("DB619_State_MPart_Write")
   "DB700_Machine_Machine{0}_StandByTime" : S5Time = PLC DB14_TP_Shortcuts.TP_Shortcuts.PageNo.1 AT %DB700.DBW24, 1 s
      on ChangeValue: SetBit("DB619_State_MPart_Write")
   "DB700_Machine_Machine{0}_StrokeCounter_KK" : Int = PLC DB14_TP_Shortcuts.TP_Shortcuts.Page_active.7 AT %DB700.DBW14, 1 s
      on ChangeValue: SetBit("DB619_State_MPart_Write")
   "DB619_State_MPart_Read" : Bool = PLC DB14_TP_Shortcuts.TP_Shortcuts.ButtonNo.6 AT %DB619.DBX6.0, 1 s
   "Machine Load Event" : Int AT %DB1.DBW0
